FUNCTION_BLOCK "Select Station PB"   // FB45, SCL
{ S7_Optimized_Access := 'TRUE' }
VERSION : 0.1
   VAR_IN_OUT
      interface : "Push Button Data";
   END_VAR
   VAR
      "Get Button Feedback" : "Push Button: State Changes";
   END_VAR
   VAR_TEMP
      _interface : "Push Button Data";
      feedback : "Push Button Data: State Change Data";
   END_VAR
BEGIN
   REGION "BUFFER IN"
       #_interface := #interface;
   END_REGION

   REGION "PROCESS USER INPUT"
       #"Get Button Feedback"(interface := #_interface,
                              state_changes := #feedback);
   END_REGION

   REGION "ANIMATIONS"
       "Select Station PB: Private: Animations"(feedback := #feedback,
                                                interface := #_interface);
   END_REGION

   REGION "BUFFER OUT"
       #interface := #_interface;
   END_REGION
END_FUNCTION_BLOCK

FUNCTION "Select Station PB: Private: Animations" : Void   // FC94, SCL
{ S7_Optimized_Access := 'TRUE' }
VERSION : 0.1
   VAR_INPUT
      feedback : "Push Button Data: State Change Data";
   END_VAR
   VAR_IN_OUT
      interface : "Push Button Data";
   END_VAR
BEGIN
   REGION "COLOR"
       #interface.animate := "Bool.Animate"(true_color := "GREEN_LIGHT_BACKGROUND",
                                             false_color := "GRAY_BACKGROUND",
                                             evaluation_signal := #feedback.actuate.actual);
   END_REGION

   REGION "VISIBILITY"
       #interface.visible := TRUE;
   END_REGION

   REGION "ENABLED STATE"
       #interface.enable := TRUE;
   END_REGION
END_FUNCTION

// folder: Display: Warehouse/002 Settings/Select WIP Button

FUNCTION_BLOCK "Select WIP PB"   // FB46, SCL
{ S7_Optimized_Access := 'TRUE' }
VERSION : 0.1
   VAR_INPUT
      settings_meta : "Setting Meta Data";
      stations : "Station: All Stations";
   END_VAR
   VAR_IN_OUT
      interface : "Push Button Data";
   END_VAR
   VAR
      "Get Button Feedback" : "Push Button: State Changes";
   END_VAR
   VAR_TEMP
      _interface : "Push Button Data";
      enable : Bool;
      feedback : "Push Button Data: State Change Data";
      visible : Bool;
   END_VAR
BEGIN
   REGION "BUFFER IN"
       #_interface := #interface;
   END_REGION

   REGION "PROCESS USER INPUT"
       #"Get Button Feedback"(interface := #_interface,
                              state_changes := #feedback);
   END_REGION

   REGION "ANIMATIONS"
       "Select WIP PB: Private: Animations"(feedback := #feedback,
                                            settings_meta := #settings_meta,
                                            stations := #stations,
                                            interface := #_interface);
   END_REGION

   REGION "BUFFER OUT"
       #interface := #_interface;
   END_REGION
END_FUNCTION_BLOCK

FUNCTION "Select WIP PB: Private: Make Visible / Enable" : Bool   // FC92, SCL
{ S7_Optimized_Access := 'TRUE' }
VERSION : 0.1
   VAR_INPUT
      settings_meta : "Setting Meta Data";
      stations : "Station: All Stations";
   END_VAR
   VAR_TEMP
      ret : Bool;
      index_of_first_selected_station : Int;
      is_hmi_station : Bool;
      first_selected_station : "Station: Single Station";
      t_select_wip : "Push Button Data";
   END_VAR
BEGIN
   REGION "ARE SELECTED STATIONS HMI STATIONS?"
       #index_of_first_selected_station := "Get First Selected Station"(#settings_meta.selected_stations.stns);
       #first_selected_station := #stations.stn[#index_of_first_selected_station];
       #is_hmi_station := "Is_HMI_Station"(#first_selected_station);
   END_REGION

   REGION "HMI STATIONS"
       IF #is_hmi_station THEN
           #ret := TRUE;
       END_IF;
   END_REGION

   REGION "RETURN"
       #"Select WIP PB: Private: Make Visible / Enable" := #ret;
   END_REGION
END_FUNCTION

FUNCTION "Select WIP PB: Private: Animations" : Void   // FC123, SCL
{ S7_Optimized_Access := 'TRUE' }
VERSION : 0.1
   VAR_INPUT
      feedback : "Push Button Data: State Change Data";
      settings_meta : "Setting Meta Data";
      stations : "Station: All Stations";
   END_VAR
   VAR_IN_OUT
      interface : "Push Button Data";
   END_VAR
BEGIN
   REGION "COLOR"
       #interface.animate := "Bool.Animate"(true_color := "GREEN_LIGHT_BACKGROUND",
                                             false_color := "GRAY_BACKGROUND",
                                             evaluation_signal := #feedback.actuate.actual);
   END_REGION

   REGION "VISIBILITY"
       #interface.visible := "Select WIP PB: Private: Make Visible / Enable"(settings_meta := #settings_meta,
                                                                              stations := #stations);
   END_REGION

   REGION "ENABLED STATE"
       #interface.enable := "Select WIP PB: Private: Make Visible / Enable"(settings_meta := #settings_meta,
                                                                             stations := #stations);
   END_REGION
END_FUNCTION

// folder: Display: Warehouse/002 Settings/Selected WIP Table

FUNCTION_BLOCK "Selected_WIP_Table"   // FB30, SCL
{ S7_Optimized_Access := 'TRUE' }
VERSION : 0.1
   VAR_INPUT
      navigation_bar : "Nav Bar Data: PLC";
      pn_library : "Recipe: PN Text Library";
      saved_wips : "Recipe: HMI Stations Saved Wips";
      settings_meta : "Setting Meta Data";
      stations : "Station: All Stations";
      wip_library : "Recipe: Wip Text Library";
   END_VAR
   VAR_IN_OUT
      stationRows : Array[0..2] of "Settings Station Row Data";
   END_VAR
   VAR
      first_selected_station : Int;
      hmi_stations_selected : Bool;
      selected_stations : Array[0.."STATION_COUNT"] of Int;
      selected_list : "Selected_WIP_Table.Selected_Array";
      row_indices : Array[0..2] of DInt;
      inst_Table_Navigation : "Table Nav";
   END_VAR
   VAR_TEMP
      i : Int;
      p_stn : Int;
      wip_code : DInt;
      visible_rows : Int;
      first_null_index : DInt;
      _hmi_saved_station_index : Int;
      _wip_index : Int;
      _wip_module : "Station: Wip: Wip Module";
   END_VAR
   // row_indices[0] := 0;
   // row_indices[1] := 1;
   // row_indices[2] := 2;
BEGIN
   REGION "CLEAR OLD CONTENTS"    
       FOR #i := 0 TO 2 DO
           #stationRows[#i].line := "Cell_Data.Hide"();
           #stationRows[#i].dropzone := "Cell_Data.Hide"();
           #stationRows[#i].wip := "Cell_Data.Hide"();
           "Button_Row.Hide_Rows"(#stationRows[#i].btnRows);
       END_FOR;
   END_REGION


   REGION "EXIT ON NO SELECTED STATION"
       IF #settings_meta.selected_stations.count = 0 THEN
           RETURN;
       END_IF;
   END_REGION


   REGION "GET ARRAY OF SELECTED STATION INDICES"
       "Array.Int.Fill"(value := "NULL_TOKEN",
                        int_array := #selected_stations);
       "Selected_Stations.Indices"(selected_stations := #settings_meta.selected_stations,
                                   selected_stations_indices := #selected_stations);
       "Selected_WIP_Table.Build_List"(selected_stations := #selected_stations,
                                       selected_wips := #settings_meta.selected_wips.wips,
                                       selected_list := #selected_list);
   END_REGION


   REGION "DETERMINE IF SELECTED STATION IS AN HMI STATION"
       #first_selected_station := "Get First Selected Station"(#settings_meta.selected_stations.stns);
       #hmi_stations_selected := "Is_HMI_Station"(#stations.stn[#first_selected_station]);
   END_REGION


   REGION "TABLE DISPLAY POINTERS"
       #first_null_index := "Selected_WIP_Table.Selected_Array.First_Occurance"(selected_array := #selected_list,
                                                                                search_term := "NULL_TOKEN");
       #inst_Table_Navigation(first_null_index := #first_null_index,
                              tblData := #selected_list.me,
                              tblDisp := #stationRows,
                              tableNav := #navigation_bar,
                              rowIndices := #row_indices);
   END_REGION


   REGION "TABLE COMPONENTS"
       #visible_rows := DINT_TO_INT(#first_null_index) - 1;
       IF #visible_rows > 2 THEN
           #visible_rows := 2;
       END_IF;
       FOR #i := 0 TO #visible_rows DO
           #p_stn := #selected_list.me[#row_indices[#i]].station_pointer;
           #wip_code := #selected_list.me[#row_indices[#i]].wip_pointer;
           #stationRows[#i].line := "Selected_WIP_Table.Line_Label.Show"(station := #stations.stn[#p_stn]);
           #stationRows[#i].dropzone := "Selected_WIP_Table.Dropzone_Label.Show"(station := #stations.stn[#p_stn]);
           #stationRows[#i].wip := "Selected_WIP_Table.Wip_Label.Show"(wip_code := #wip_code,
                                                                       wip_library := #wip_library);
           #_wip_module := "Selected_WIP_Table.Get_WIP_Module"(stations := #stations,
                                                               saved_wips := #saved_wips,
                                                               station_pointer := #p_stn,
                                                               wip_code := #wip_code);
           "Button_Row.Show_Rows"(selected_butttons := #settings_meta.selected_btns,
                                  wip_module := #_wip_module,
                                  pn_library := #pn_library,
                                  button_rows := #stationRows[#i].btnRows);
       END_FOR;
   END_REGION
END_FUNCTION_BLOCK

FUNCTION "Selected_WIP_Table.Build_List" : Void   // FC219, SCL
{ S7_Optimized_Access := 'TRUE' }
VERSION : 0.1
   VAR_INPUT
      selected_stations : Array[*] of Int;
      selected_wips : Array[*] of DInt;
   END_VAR
   VAR_IN_OUT
      selected_list : "Selected_WIP_Table.Selected_Array";
   END_VAR
   VAR_TEMP
      _i : DInt;
      _j : DInt;
      _length : Struct
         stations : DInt;
         wips : DInt;
      END_STRUCT;
      _p : DInt;
   END_VAR
BEGIN
   REGION "PREPARE ARRAY"
       "Selected_WIP_Table.Selected_Array.Fill"(token := -1,
                                                selected_list := #selected_list);
   END_REGION


   REGION "GET UPPER LIMIT FOR OUTER LOOP"
       #_length.stations := "Array.Int.First_Occurance"(int_array := #selected_stations,
                                                        search_term := "NULL_TOKEN");
       #_length.stations -= 1;
       #_length.stations := "DInt.Clip.Minimum"(value := #_length.stations,
                                                minimum := 0);
   END_REGION


   REGION "GET LIMIT FOR INNER LOOP"
       #_length.wips := "Array.DInt.First_Occurance"(dint_array := #selected_wips,
                                                     search_term := "NULL_TOKEN");
       #_length.wips -= 1;
       #_length.wips := "DInt.Clip.Minimum"(value := #_length.wips,
                                            minimum := 0);
   END_REGION


   REGION "BUILD ARRAY"
       FOR #_i := 0 TO #_length.stations DO
           FOR #_j := 0 TO #_length.wips DO
               #_p := #_i * (#_length.wips + 1) + #_j;
               #selected_list.me[#_p].station_pointer := #selected_stations[#_i];
               #selected_list.me[#_p].wip_pointer := #selected_wips[#_j];
           END_FOR;
       END_FOR;
   END_REGION
END_FUNCTION

FUNCTION "Selected_WIP_Table.Selected_Array.Fill" : Void   // FC221, SCL
{ S7_Optimized_Access := 'TRUE' }
VERSION : 0.1
   VAR_INPUT
      token : Int;
   END_VAR
   VAR_IN_OUT
      selected_list : "Selected_WIP_Table.Selected_Array";
   END_VAR
   VAR_TEMP
      _i : DInt;
      _length : DInt;
   END_VAR
BEGIN
   #_length := UDINT_TO_DINT("Array.Any.Length"(#selected_list.me));
   #_length -= 1;

   FOR #_i := 0 TO #_length DO
       #selected_list.me[#_i].station_pointer := #token;
       #selected_list.me[#_i].wip_pointer := INT_TO_DINT(#token);
   END_FOR;
END_FUNCTION

FUNCTION "Selected_WIP_Table.Selected_Array.Is_Element" : Bool   // FC228, SCL
{ S7_Optimized_Access := 'TRUE' }
VERSION : 0.1
   VAR_INPUT
      selected_array : "Selected_WIP_Table.Selected_Array";
      search_term : Int;
   END_VAR
   VAR_TEMP
      _i : DInt;
      _length : DInt;
   END_VAR
BEGIN
   REGION "LOCAL VARIABLES"
       #_length := UDINT_TO_DINT("Array.Any.Length"(#selected_array.me)) - 1;
   END_REGION


   REGION "SEARCH ARRAY"
       FOR #_i := 0 TO #_length DO
           IF #selected_array.me[#_i].station_pointer <> #search_term THEN
               CONTINUE;
           END_IF;
           #"Selected_WIP_Table.Selected_Array.Is_Element" := TRUE;
           RETURN;
       END_FOR;
   END_REGION


   REGION "NOT FOUND"
       #"Selected_WIP_Table.Selected_Array.Is_Element" := FALSE;
       RETURN;
   END_REGION
END_FUNCTION

FUNCTION "Selected_WIP_Table.Selected_Array.First_Occurance" : DInt   // FC229, SCL
{ S7_Optimized_Access := 'TRUE' }
VERSION : 0.1
   VAR_INPUT
      selected_array : "Selected_WIP_Table.Selected_Array";
      search_term : Int;
   END_VAR
   VAR_TEMP
      _i : DInt;
      _length : UDInt;
   END_VAR
BEGIN
   REGION "NOTES"
       (* 
       This function returns the first occurance of the search term.
       This function meant for use with collapsed arrays.
       See "Array.Int.Collapse" for collapse functionality.
       *)
   END_REGION


   REGION "GET LENGTH OF INPUT ARRAY"
       #_length := "Array.Any.Length"(#selected_array.me);
   END_REGION


   REGION "FIND FIRST SEARCH TERM, -1 IF NONE"
       (*
       Its worth noting that "Array.Int.Is_Element" could return the index of the search term
       as an output, saving the processor some work. 
       The rework is justified by increased encapsulation.
       The time complexity for "Array.Int.First_Occurance" remains O(n).
       *)
       IF NOT "Selected_WIP_Table.Selected_Array.Is_Element"(selected_array:=#selected_array, search_term:=#search_term) THEN
           #"Selected_WIP_Table.Selected_Array.First_Occurance" := -1;
           RETURN;
       END_IF;
       WHILE #selected_array.me[#_i].station_pointer <> #search_term AND DINT_TO_UDINT(#_i) < #_length DO
           #_i += 1;
       END_WHILE;
   END_REGION


   REGION "SEARCH TERM FOUND"
       #"Selected_WIP_Table.Selected_Array.First_Occurance" := #_i;
       RETURN;
   END_REGION
END_FUNCTION

FUNCTION "Selected_WIP_Table.Get_WIP_Module" : "Station: Wip: Wip Module"   // FC234, SCL
{ S7_Optimized_Access := 'TRUE' }
VERSION : 0.1
   VAR_INPUT
      stations : "Station: All Stations";
      saved_wips : "Recipe: HMI Stations Saved Wips";
      station_pointer : Int;
      wip_code : DInt;
   END_VAR
   VAR_TEMP
      _hmi_station_pointer : Int;
      _wip_pointer : Int;
   END_VAR
BEGIN
   IF #wip_code = "NULL_TOKEN" THEN
       #"Selected_WIP_Table.Get_WIP_Module" := #stations.stn[#station_pointer].wipCmpts;
       RETURN;
   END_IF;

   #_hmi_station_pointer := "WIP.Global_Index_to_HMI_Station_Index"(global_index := #station_pointer,
                                                                    saved_WIPs := #saved_wips);

   #_wip_pointer := "WIP.Code_to_Index"(saved_wip := #saved_wips.stn[#_hmi_station_pointer],
                                        wip_code := #wip_code);

   #"Selected_WIP_Table.Get_WIP_Module" := #saved_wips.stn[#_hmi_station_pointer].wip[#_wip_pointer];
   RETURN;
END_FUNCTION

// folder: Display: Warehouse/002 Settings/Selected WIP Table/Button Row

FUNCTION "Button_Row.Hide" : "Settings Station Row Button Row Data"   // FC210, SCL
{ S7_Optimized_Access := 'TRUE' }
VERSION : 0.1
   VAR_TEMP
      _ret : "Settings Station Row Button Row Data";
   END_VAR
BEGIN
   #_ret.button := "Cell_Data.Hide"();
   #_ret.total := "Cell_Data.Hide"();
   #_ret.critical := "Cell_Data.Hide"();
   #_ret.singlePN := "Cell_Data.Hide"();
   #_ret.doublePN := "Cell_Data.Hide"();
   #"Button_Row.Hide" := #_ret;
END_FUNCTION

FUNCTION "Button_Row.Hide_Rows" : Void   // FC211, SCL
{ S7_Optimized_Access := 'TRUE' }
VERSION : 0.1
   VAR_IN_OUT
      button_rows : Array[*] of "Settings Station Row Button Row Data";
   END_VAR
   VAR_TEMP
      _i : Int;
   END_VAR
BEGIN
   FOR #_i := 0 TO UDINT_TO_INT("Array.Any.Length"(#button_rows)) - 1 DO
       #button_rows[#_i] := "Button_Row.Hide"();
   END_FOR;
END_FUNCTION

FUNCTION "Button_Row.Show" : "Settings Station Row Button Row Data"   // FC212, SCL
{ S7_Optimized_Access := 'TRUE' }
VERSION : 0.1
   VAR_INPUT
      button_number : Int;
      selected : Bool;
      pn_library : "Recipe: PN Text Library";
      wip_module : "Station: Wip: Wip Module";
   END_VAR
   VAR_TEMP
      _return : "Settings Station Row Button Row Data";
      _pn : "Cell Data";
   END_VAR
BEGIN
   #_return.button := "Button_Row.Button_Label.Show"(button_number := #button_number,
                                                     selected := #selected);

   #_return.total := "Button_Row.Total.Show"(selected := #selected,
                                             button_number := #button_number,
                                             wip_module := #wip_module);

   #_return.critical := "Button_Row.Critical.Show"(button_number := #button_number,
                                                   selected := #selected,
                                                   wip_module := #wip_module);

   #_pn := "Button_Row.Part_Number.Show"(button_number := #button_number,
                                         pn_library := #pn_library,
                                         selected := #selected,
                                         wip_module := #wip_module);

   IF "Part_Number.Is_Single"(#wip_module.pnCode[#button_number]) THEN
       #_return.singlePN := #_pn;
   END_IF;
   IF "Part_Number.Is_Double"(#wip_module.pnCode[#button_number]) THEN
       #_return.doublePN := #_pn;
   END_IF;
   #"Button_Row.Show" := #_return;
END_FUNCTION

FUNCTION "Button_Row.Show_Rows" : Void   // FC218, SCL
{ S7_Optimized_Access := 'TRUE' }
VERSION : 0.1
   VAR_INPUT
      selected_butttons : "Selected Buttons";
      wip_module : "Station: Wip: Wip Module";
      pn_library : "Recipe: PN Text Library";
   END_VAR
   VAR_IN_OUT
      button_rows : Array[*] of "Settings Station Row Button Row Data";
   END_VAR
   VAR_TEMP
      _i : Int;
      _remap : Int;
   END_VAR
BEGIN
   FOR #_i := 0 TO UDINT_TO_INT("Array.Any.Length"(#button_rows)) - 1 DO
       #_remap := "KP8.DURL_to_LRUD"(#_i);
       #button_rows[#_i] := "Button_Row.Show"(button_number := #_remap,
                                              selected := #selected_butttons.btns[#_i],
                                              pn_library := #pn_library,
                                              wip_module := #wip_module);
   END_FOR;
END_FUNCTION

// folder: Display: Warehouse/002 Settings/Selected WIP Table/Button Row/Single Button

FUNCTION "Button_Row.Button_Label.Show" : "Cell Data"   // FC213, SCL
{ S7_Optimized_Access := 'TRUE' }
VERSION : 0.1
   VAR_INPUT
      button_number : Int;
      selected : Bool;
   END_VAR
   VAR_TEMP
      _animate : Int;
      _data : WString;
   END_VAR
BEGIN
   #_animate := "Bool.Animate"(true_color := "BLUE_LIGHT_BACKGROUND",
                               false_color := "GRAY_BACKGROUND",
                               evaluation_signal := #selected);
   #_data := "Trim"("Strip Sign"(INT_TO_WSTRING(#button_number)));
   #"Button_Row.Button_Label.Show" := "Cell_Data.Show"(animate := #_animate, data := #_data);
END_FUNCTION

FUNCTION "Button_Row.Total.Show" : "Cell Data"   // FC214, SCL
{ S7_Optimized_Access := 'TRUE' }
VERSION : 0.1
   VAR_INPUT
      button_number : Int;
      selected : Bool;
      wip_module : "Station: Wip: Wip Module";
   END_VAR
   VAR_TEMP
      _animation : Int;
      _data : WString;
   END_VAR
BEGIN
   #_animation := "Bool.Animate"(true_color := "BLUE_LIGHT_BACKGROUND",
                                 false_color := "GRAY_BACKGROUND",
                                 evaluation_signal := #selected);

   #_data := "Button_Row.Total.Extract_String"(button_number := #button_number,
                                               wip_module := #wip_module);

   #"Button_Row.Total.Show" := "Cell_Data.Show"(animate := #_animation,
                                                data := #_data);
END_FUNCTION

FUNCTION "Button_Row.Critical.Show" : "Cell Data"   // FC215, SCL
{ S7_Optimized_Access := 'TRUE' }
VERSION : 0.1
   VAR_INPUT
      button_number : Int;
      selected : Bool;
      wip_module : "Station: Wip: Wip Module";
   END_VAR
   VAR_TEMP
      _animate : Int;
      _data : WString;
   END_VAR
BEGIN
   #_animate := "Bool.Animate"(true_color := "BLUE_LIGHT_BACKGROUND",
                               false_color := "GRAY_BACKGROUND",
                               evaluation_signal := #selected);

   #_data := "Button_Row.Critical.Extract_String"(button_number := #button_number,
                                                  wip_module := #wip_module);

   #"Button_Row.Critical.Show" := "Cell_Data.Show"(animate := #_animate, data := #_data);
END_FUNCTION

FUNCTION "Button_Row.Part_Number.Show" : "Cell Data"   // FC217, SCL
{ S7_Optimized_Access := 'TRUE' }
VERSION : 0.1
   VAR_INPUT
      button_number : Int;
      pn_library : "Recipe: PN Text Library";
      selected : Bool;
      wip_module : "Station: Wip: Wip Module";
   END_VAR
   VAR_TEMP
      _animation : Int;
      _data : WString;
      _pn_code : DInt;
   END_VAR
BEGIN
   #_animation := "Bool.Animate"(true_color := "BLUE_LIGHT_BACKGROUND",
                                 false_color := "GRAY_BACKGROUND",
                                 evaluation_signal := #selected);

   #_pn_code := "Button_Row.Part_Number.Extract_Code"(button_number := #button_number,
                                                      wip_module := #wip_module);

   #_data := "Part_Number.Code_to_WString"(pnLib := #pn_library,
                                           pnCode := #_pn_code);

   #"Button_Row.Part_Number.Show" := "Cell_Data.Show"(animate := #_animation,
                                                      data := #_data);
END_FUNCTION

FUNCTION "Button_Row.Total.Extract_String" : WString   // FC230, SCL
{ S7_Optimized_Access := 'TRUE' }
VERSION : 0.1
   VAR_INPUT
      button_number : Int;
      wip_module : "Station: Wip: Wip Module";
   END_VAR
BEGIN
   #"Button_Row.Total.Extract_String" := "Timer.Real_to_WString"(#wip_module.timers.ptAllotted[#button_number]);
   RETURN;
END_FUNCTION

FUNCTION "Button_Row.Part_Number.Extract_Code" : DInt   // FC231, SCL
{ S7_Optimized_Access := 'TRUE' }
VERSION : 0.1
   VAR_INPUT
      button_number : Int;
      wip_module : "Station: Wip: Wip Module";
   END_VAR
   VAR_TEMP
      _hmi_station_pointer : Int;
      _pn_code : DInt;
      _wip_pointer : Int;
   END_VAR
BEGIN
   #"Button_Row.Part_Number.Extract_Code" := #wip_module.pnCode[#button_number];
   RETURN;
END_FUNCTION

FUNCTION "Button_Row.Critical.Extract_String" : WString   // FC232, SCL
{ S7_Optimized_Access := 'TRUE' }
VERSION : 0.1
   VAR_INPUT
      button_number : Int;
      wip_module : "Station: Wip: Wip Module";
   END_VAR
BEGIN
   #"Button_Row.Critical.Extract_String" := "Timer.Real_to_WString"(#wip_module.timers.ptCritical[#button_number]);
   RETURN;
END_FUNCTION

// folder: Display: Warehouse/002 Settings/Selected WIP Table/Dropzone Label

FUNCTION "Selected_WIP_Table.Dropzone_Label.Show" : "Cell Data"   // FC200, SCL
{ S7_Optimized_Access := 'TRUE' }
VERSION : 0.1
   VAR_INPUT
      station : "Station: Single Station";
   END_VAR
BEGIN
   #"Selected_WIP_Table.Dropzone_Label.Show" := "Cell_Data.Show"(animate := "GRAY_BACKGROUND",
                                                                 data := "Trim"("Strip Sign"(USINT_TO_WSTRING(#station.id.dropZone))));
END_FUNCTION

// folder: Display: Warehouse/002 Settings/Selected WIP Table/Line Label

FUNCTION "Selected_WIP_Table.Line_Label.Show" : "Cell Data"   // FC199, SCL
{ S7_Optimized_Access := 'TRUE' }
VERSION : 0.1
   VAR_INPUT
      station : "Station: Single Station";
   END_VAR
   VAR CONSTANT
      SHOW : Bool := TRUE;
   END_VAR
BEGIN
   #"Selected_WIP_Table.Line_Label.Show" := "Cell_Data.Show"(animate := "GRAY_BACKGROUND",
                                                             data := #station.id.lineName);
END_FUNCTION

// folder: Display: Warehouse/002 Settings/Selected WIP Table/Wip Label

FUNCTION "Selected_WIP_Table.Wip_Label.Show" : "Cell Data"   // FC201, SCL
{ S7_Optimized_Access := 'TRUE' }
VERSION : 0.1
   VAR_INPUT
      wip_code : DInt;
      wip_library : "Recipe: Wip Text Library";
   END_VAR
   VAR_TEMP
      _delimeters : Array[0..9] of WString[1];
      _data : WString;
   END_VAR
   VAR CONSTANT
      SHOW : Bool := TRUE;
   END_VAR
BEGIN
   IF #wip_code = "NULL_TOKEN" THEN
       #"Selected_WIP_Table.Wip_Label.Show" := "Cell_Data.Hide"();
       RETURN;
   END_IF;

   #_data := "WIP.Code_to_WString"(wipTxtLib := #wip_library,
                                   code := #wip_code);
   #_delimeters[0] := WSTRING#' ';
   #_delimeters[1] := WSTRING#'-';
   #_delimeters[2] := WSTRING#'.';
   #_data := "WString.Word_Wrap"(delimeters := #_delimeters,
                                 line_length := 20,
                                 wstring_in := #_data);

   #"Selected_WIP_Table.Wip_Label.Show" := "Cell_Data.Show"(animate := "GRAY_BACKGROUND", data := #_data);
END_FUNCTION

// folder: Display: Warehouse/002 Settings/Total IO Field

FUNCTION_BLOCK "Total_IO_Field"   // FB49, SCL
{ S7_Optimized_Access := 'TRUE' }
VERSION : 0.1
   VAR_INPUT
      settings_meta : "Setting Meta Data";
      stations : "Station: All Stations";
   END_VAR
   VAR_IN_OUT
      interface : "IO Field Data: Label with Data";
      state_changes : "State Changes: Real";
   END_VAR
   VAR
      Total_IO_Field : "IO Field: State Changes";
      Detect_State_Changes : "Real.State_Change";
   END_VAR
   VAR_TEMP
      _interface : "IO Field Data: Label with Data";
      feedback : "IO Field: State Change Data";
   END_VAR
BEGIN
   REGION "BUFFER IN"
       #_interface := #interface;
   END_REGION

   REGION "PROCESS USER INPUT"
       #Total_IO_Field(interface := #_interface,
                       feedback := #feedback);
       #Detect_State_Changes(value := "Timer.WString_to_Real"(#interface.value),
                             get_real := #state_changes);
   END_REGION

   REGION "BUFFER OUT"
       "Total_IO_Field.Animate"(feedback := #feedback,
                                settings_meta := #settings_meta,
                                stations := #stations,
                                interface := #_interface);
   END_REGION

   REGION "BUFFER OUT"
       #interface := #_interface;
   END_REGION
END_FUNCTION_BLOCK

FUNCTION "Total_IO_Field.Make_Visible_Enable" : Bool   // FC189, SCL
{ S7_Optimized_Access := 'TRUE' }
VERSION : 0.1
   VAR_INPUT
      setting_meta : "Setting Meta Data";
   END_VAR
BEGIN
   #"Total_IO_Field.Make_Visible_Enable" := #setting_meta.selected_btns.count > 0;
END_FUNCTION

FUNCTION "Total_IO_Field.Animate" : Void   // FC190, SCL
{ S7_Optimized_Access := 'TRUE' }
VERSION : 0.1
   VAR_INPUT
      feedback : "IO Field: State Change Data";
      settings_meta : "Setting Meta Data";
      stations : "Station: All Stations";
   END_VAR
   VAR_IN_OUT
      interface : "IO Field Data: Label with Data";
   END_VAR
   VAR_TEMP
      _visible_enabled : Bool;
   END_VAR
BEGIN
   REGION "COLOR"
   #interface.animate := "WHITE_BACKGROUND";
   END_REGION


   REGION "SET STATE"
       #_visible_enabled := "Total_IO_Field.Make_Visible_Enable"(setting_meta := #settings_meta);
   END_REGION


   REGION "VISIBILITY
       #interface.visible := #_visible_enabled;
   END_REGION


   REGION "ENABLE"
       #interface.enable := #_visible_enabled;
   END_REGION


   REGION "POPULATE VALUE"
       IF #settings_meta.button_selection_change.selection_change THEN
           #interface.value := "Total_IO_Field.Populate_Value"(hidden := NOT #_visible_enabled,
                                                               selected_buttons := #settings_meta.selected_btns,
                                                               selected_stations := #settings_meta.selected_stations,
                                                               stations := #stations);
       END_IF;
   END_REGION
END_FUNCTION

FUNCTION "Total_IO_Field.Populate_Value" : WString   // FC292, SCL
{ S7_Optimized_Access := 'TRUE' }
VERSION : 0.1
   VAR_INPUT
      hidden : Bool;
      selected_buttons : "Selected Buttons";
      selected_stations : "Selected Stations";
      stations : "Station: All Stations";
   END_VAR
   VAR_TEMP
      _critical : WString;
      _p_station : Int;
      _p_button : Int;
   END_VAR
   VAR CONSTANT
      BLANK : WString;
      ZERO : WChar := WCHAR#'0';
   END_VAR
BEGIN
   IF #hidden THEN
       #"Total_IO_Field.Populate_Value" := #BLANK;
       RETURN;
   END_IF;
   #_p_station := "Selected_Stations.Get_First_Selected_Station"(#selected_stations);
   #_p_button := "Selected_Buttons.Get_First_Selected_Button"(#selected_buttons);
   #_critical := "Timer.Real_to_WString"(#stations.stn[#_p_station].wipCmpts.timers.ptAllotted[#_p_button]);
   #"Total_IO_Field.Populate_Value" := #_critical;
END_FUNCTION

// folder: Display: Warehouse/Pop Ups/Pop Up Utilities

FUNCTION "Animate Array: PB Data Activation" : Bool   // FC95, SCL
{ S7_Optimized_Access := 'TRUE' }
VERSION : 0.1
   VAR_INPUT
      element_index : Int;
      visible_element_count : Int;
   END_VAR
   VAR_TEMP
      ret : Bool;
   END_VAR
BEGIN
   REGION "TURN ON A NUMBER OF BUTTONS EQUAL TO THE NUMBER OF STATIONS"
       IF #element_index < #visible_element_count THEN
           #ret := TRUE;
       END_IF;
       IF #element_index >= #visible_element_count THEN
           #ret := FALSE;
       END_IF;
   END_REGION

   REGION "RETURN"
       #"Animate Array: PB Data Activation" := #ret;
   END_REGION
END_FUNCTION

FUNCTION "Pop Up: Nav Bar: Button Animation" : Void   // FC97, SCL
{ S7_Optimized_Access := 'TRUE' }
VERSION : 0.1
   VAR_INPUT
      selectable_elements : Int;
      visible_rows : Int;
   END_VAR
   VAR_IN_OUT
      button : "Push Button Data";
   END_VAR
   VAR_TEMP
      ret : "Push Button Data";
   END_VAR
BEGIN
   REGION "SHOW NAV BAR"
       IF #selectable_elements > #visible_rows THEN

           REGION "GET CURRENT STATE FOR PRESS"
               #ret := #button;
           END_REGION

           REGION "ANIMATION"
               #ret.animate := "Bool.Animate"(true_color := "GREEN_LIGHT_BACKGROUND",
                                              false_color := "GRAY_BACKGROUND",
                                              evaluation_signal := #button.actuate);
           END_REGION

           REGION "ENABLE"
               #ret.enable := TRUE;
           END_REGION

           REGION "LIST SELECT"
               #ret.listSelect := 0;
           END_REGION

           REGION "VISIBLE"
               #ret.visible := TRUE;
           END_REGION

       END_IF;
   END_REGION


   REGION "HIDE NAV BAR"
       IF #selectable_elements <= #visible_rows THEN

           REGION "DIABLE"
               #ret.enable := FALSE;
           END_REGION

           REGION "INVISIBLE"
               #ret.visible := FALSE;
           END_REGION

       END_IF;
   END_REGION


   REGION "RETURN"
       #button := #ret;
   END_REGION
END_FUNCTION

FUNCTION "Pop Up: Map Select Button Actuations" : Void   // FC117, SCL
{ S7_Optimized_Access := 'TRUE' }
VERSION : 0.1
   VAR_INPUT
      screen_elements : Variant;
   END_VAR
   VAR_IN_OUT
      actuations_as_ints : Variant;
   END_VAR
   VAR_TEMP
      i : Int;
      len_udint : UDInt;
      len_int : Int;
      ret : Array[0..#u_bound_simple] of Int;
      status : Int;
      t_select_btns : Array[0..#u_bound_complex] of "Push Button Data";
   END_VAR
   VAR CONSTANT
      u_bound_simple : Int := 99;
      u_bound_complex : Int := 29;
   END_VAR
BEGIN
   REGION "GET PARAMETERS"
       #len_udint := CountOfElements(#screen_elements);
       #len_int := UDINT_TO_INT(#len_udint) - 1;
   END_REGION

   REGION "COPY TO LOCAL"
       #status := MOVE_BLK_VARIANT(SRC := #screen_elements,
                                   COUNT := #len_udint,
                                   SRC_INDEX := 0,
                                   DEST_INDEX := 0,
                                   DEST => #t_select_btns);
   END_REGION

   REGION "MAP ACTUATIONS"    
       FOR #i := 0 TO #len_int DO
           IF #t_select_btns[#i].actuate THEN
               #ret[#i] := 1;
           END_IF;
       END_FOR;
   END_REGION

   REGION "RETURN"
       #status := MOVE_BLK_VARIANT(SRC := #ret,
                                   COUNT := #len_udint,
                                   SRC_INDEX := 0,
                                   DEST_INDEX := 0,
                                   DEST => #actuations_as_ints);
   END_REGION
END_FUNCTION

FUNCTION "Pop Up: Nav Bar: Animate" : Void   // FC135, SCL
{ S7_Optimized_Access := 'TRUE' }
VERSION : 0.1
   VAR_INPUT
      selectable_element_count : Int;
      visible_rows : Int;
   END_VAR
   VAR_IN_OUT
      nav_bar : "Nav Bar Data";
   END_VAR
BEGIN
       REGION "NOTES"
           // mapping is necessary because hmi faceplate data structures
           // cannot consist of embedded udts
       END_REGION

       REGION "MAP HMI TO PLC"
           "NavBar: Map HMI to PLC"(hmi := #nav_bar.hmi,
                                          plc := #nav_bar.plc);
       END_REGION

       REGION "ANIMATION CALLS"
           "Pop Up: Nav Bar: Button Animation"(selectable_elements := #selectable_element_count,
                                               visible_rows := #visible_rows,
                                               button := #nav_bar.plc.top);
           "Pop Up: Nav Bar: Button Animation"(selectable_elements := #selectable_element_count,
                                               visible_rows := #visible_rows,
                                               button := #nav_bar.plc.pageUp);
           "Pop Up: Nav Bar: Button Animation"(selectable_elements := #selectable_element_count,
                                               visible_rows := #visible_rows,
                                               button := #nav_bar.plc.lineUp);
           "Pop Up: Nav Bar: Button Animation"(selectable_elements := #selectable_element_count,
                                               visible_rows := #visible_rows,
                                               button := #nav_bar.plc.lineDown);
           "Pop Up: Nav Bar: Button Animation"(selectable_elements := #selectable_element_count,
                                               visible_rows := #visible_rows,
                                               button := #nav_bar.plc.pageDown);
           "Pop Up: Nav Bar: Button Animation"(selectable_elements := #selectable_element_count,
                                               visible_rows := #visible_rows,
                                               button := #nav_bar.plc.bottom);
       END_REGION

       REGION "MAP PLC TO HMI"
           "NavBar: Map PLC to HMI"(plc := #nav_bar.plc,
                                          hmi := #nav_bar.hmi);
       END_REGION
END_FUNCTION

FUNCTION "Clear WIP Selection Meta Data" : Void   // FC193, SCL
{ S7_Optimized_Access := 'TRUE' }
VERSION : 0.1
   VAR_IN_OUT
      selected_wips : "Selected Wips";
   END_VAR
   VAR_TEMP
      i : Int;
      selected_wips_array : Array[0.."WIP_COUNT"] of DInt;
   END_VAR
BEGIN
   "Array.DInt.Fill"(int_in := INT_TO_DINT("NULL_TOKEN"),
                     array_out => #selected_wips.wips);
   #selected_wips.count := 0;
END_FUNCTION

FUNCTION "Clear Button Selection Meta Data" : Void   // FC194, SCL
{ S7_Optimized_Access := 'TRUE' }
VERSION : 0.1
   VAR_IN_OUT
      selected_buttons : "Selected Buttons";
   END_VAR
   VAR_TEMP
      i : Int;
   END_VAR
BEGIN
   #selected_buttons.count := 0;
   FOR #i := 0 TO "BUTTON_COUNT" DO
       #selected_buttons.btns[#i] := FALSE;
   END_FOR;
END_FUNCTION

// folder: Display: Warehouse/Pop Ups/Select Buttons

FUNCTION_BLOCK "Pop Up: Select Buttons"   // FB25, SCL
{ S7_Optimized_Access := 'TRUE' }
VERSION : 0.1
   VAR_IN_OUT
      interface : "Select Button";
      selected_buttons : "Selected Buttons";
      meta_data : "Setting Meta Data";
   END_VAR
   VAR
      "inst Pop Up: Select Buttons: Select Buttons" : "Pop Up: Select Buttons: Select Buttons";
      Button_Selection_Change : "Selected_Buttons.Selection_Change";
   END_VAR
BEGIN
   REGION "ANIMATION"
       "Pop Up: Select Buttons: Animations"(interface := #interface,
                                            selected := #selected_buttons);
   END_REGION


   REGION "PERFORM BUTTON SELECTION"
       #"inst Pop Up: Select Buttons: Select Buttons"(interface := #interface,
                                                      selected_buttons := #selected_buttons);
   END_REGION


   REGION "CHECK FOR BUTTON SELECTION CHANGE"
       #Button_Selection_Change(selected_buttons := #selected_buttons,
                                selection_change := #meta_data.button_selection_change);
   END_REGION


   REGION "HOUSE KEEPING FOR STATION SELECTION CHANGE"
       IF #meta_data.station_selection_change.selection_change THEN
           "Clear Button Selection Meta Data"(#meta_data.selected_btns);
       END_IF;
   END_REGION
END_FUNCTION_BLOCK

FUNCTION_BLOCK "Pop Up: Select Buttons: Select Buttons"   // FB27, SCL
{ S7_Optimized_Access := 'TRUE' }
VERSION : 0.1
   VAR_IN_OUT
      interface : "Select Button";
      selected_buttons : "Selected Buttons";
   END_VAR
   VAR
      "inst Pulses: Button Collection" : "Pulses: Button Collection";
   END_VAR
   VAR_TEMP
      actuation_pulses : Array[0.."BUTTON_COUNT"] of Bool;
      actuations_as_ints : Array[0.."BUTTON_COUNT"] of Int;
      i : Int;
      pulses_as_ints : Array[0.."BUTTON_COUNT"] of Int;
   END_VAR
BEGIN
   "Pop Up: Map Select Button Actuations"(screen_elements := #interface.buttons,
                                          actuations_as_ints := #actuations_as_ints);
   #"inst Pulses: Button Collection"(btns := #actuations_as_ints,
                                     pulses := #pulses_as_ints);
   "Pop Up: Select Buttons: Pulse Ints to Bools"(pulses_as_ints := #pulses_as_ints,
                                                 pulses_as_bools => #actuation_pulses);
   FOR #i := 0 TO "BUTTON_COUNT" DO
       "Toggle"(pulse := #actuation_pulses[#i],
                state := #selected_buttons.btns[#i]);
   END_FOR;
   #selected_buttons.count := "Count Selected Buttons"(#selected_buttons.btns);
END_FUNCTION_BLOCK

FUNCTION_BLOCK "Selected_Buttons.Selection_Change"   // FB59, SCL
{ S7_Optimized_Access := 'TRUE' }
VERSION : 0.1
   VAR_INPUT
      selected_buttons : "Selected Buttons";
   END_VAR
   VAR_IN_OUT
      selection_change : "Selected_Buttons.Selection_Change.UDT";
   END_VAR
   VAR
      old : Struct
         selected_buttons : "Selected Buttons";
      END_STRUCT;
   END_VAR
   VAR_TEMP
      _i : Int;
      _return : "Selected_Buttons.Selection_Change.UDT";
   END_VAR
BEGIN
   REGION "SCAN FOR CHANGE"
       FOR #_i := 0 TO "BUTTON_COUNT" DO
           IF #selected_buttons.btns[#_i] <> #old.selected_buttons.btns[#_i] THEN
               #_return.selection_change := TRUE;
               #_return.button_index := #_i;
               IF #selected_buttons.btns[#_i] AND NOT #old.selected_buttons.btns[#_i] THEN
                   #_return.rising := TRUE;
                   #_return.falling := FALSE;
               END_IF;
               IF NOT #selected_buttons.btns[#_i] AND #old.selected_buttons.btns[#_i] THEN
                   #_return.rising := FALSE;
                   #_return.falling := TRUE;
               END_IF;
               EXIT;
           END_IF;
       END_FOR;
   END_REGION


   REGION "SAVE TO OLD"
       #old.selected_buttons := #selected_buttons;
   END_REGION


   REGION "RETURN"
       #selection_change := #_return;
   END_REGION
END_FUNCTION_BLOCK

FUNCTION "Pop Up: Select Buttons: Animations" : Void   // FC116, SCL
{ S7_Optimized_Access := 'TRUE' }
VERSION : 0.1
   VAR_IN_OUT
      interface : "Select Button";
      selected : "Selected Buttons";
   END_VAR
   VAR_TEMP
      i : Int;
      selected_stations_count : Int;
      t_interface : "Select Button";
   END_VAR
BEGIN
   REGION "COPY TO LOCAL"
       #t_interface := #interface;
   END_REGION

   REGION "CLOSE POPUP BUTTON"
       #t_interface.close_screen.animate := "Bool.Animate"(true_color := "GREEN_LIGHT_BACKGROUND",
                                                           false_color := "RED_LIGHT_BACKGROUND",
                                                           evaluation_signal := #interface.close_screen.actuate);
   END_REGION


   REGION "BUTTON SELECTION BUTTONS"
       FOR #i := 0 TO "BUTTON_COUNT" DO
           #t_interface.buttons[#i].animate := "Bool.Animate"(true_color := "GREEN_LIGHT_BACKGROUND",
                                                              false_color := "GRAY_BACKGROUND",
                                                              evaluation_signal := #interface.buttons[#i].actuate);
           #t_interface.buttons[#i].enable := TRUE;
           #t_interface.buttons[#i].visible := TRUE;
           IF #selected.btns[#i] THEN
               #t_interface.buttons[#i].animate := "BLUE_LIGHT_BACKGROUND";
           END_IF;
       END_FOR;
   END_REGION


   REGION "DRAW"
       #interface := #t_interface;
   END_REGION
END_FUNCTION

FUNCTION "Pop Up: Select Buttons: Pulse Ints to Bools" : Void   // FC118, SCL
{ S7_Optimized_Access := 'TRUE' }
VERSION : 0.1
   VAR_INPUT
      pulses_as_ints : Array[0.."BUTTON_COUNT"] of Int;
   END_VAR
   VAR_OUTPUT
      pulses_as_bools : Array[0.."BUTTON_COUNT"] of Bool;
   END_VAR
   VAR_TEMP
      i : Int;
      ret : Array[0.."BUTTON_COUNT"] of Bool;
   END_VAR
BEGIN
   REGION "MAP TO BOOLS"
       FOR #i := 0 TO "BUTTON_COUNT" DO
           #ret[#i] := #pulses_as_ints[#i].%X0;
       END_FOR;
   END_REGION

   REGION "RETURN"
       #pulses_as_bools := #ret;
   END_REGION
END_FUNCTION

// folder: Display: Warehouse/Pop Ups/Select Station

FUNCTION_BLOCK "Pop Up: Select Stations"   // FB21, SCL
{ S7_Optimized_Access := 'TRUE' }
VERSION : 0.1
   VAR_INPUT
      all_stations : "Station: All Stations";
      saved_WIPs : "Recipe: HMI Stations Saved Wips";
   END_VAR
   VAR_IN_OUT
      interface : "Select Station";
      meta_data : "Setting Meta Data";
   END_VAR
   VAR
      "inst Patch for Table Nav in Select Station Popup" : "Patch for Table Nav in Select Station Popup";
      "inst Select Station Button Pulses" : "Pulses: Button Collection";
      "inst Selection Change" : "Selected_Stations.Selection_Change";
      "inst Table Nav" : "Table Nav";
      vis_stns_as_dint : Array[0.."_SELECT_STATION_BUTTON_COUNT"] of DInt;
      visable_stns : Array[0.."_SELECT_STATION_BUTTON_COUNT"] of Int;
   END_VAR
   VAR_TEMP
      actuations_as_ints : Array[0.."_SELECT_STATION_BUTTON_COUNT"] of Int;
      actuation_pulses : Array[0.."_SELECT_STATION_BUTTON_COUNT"] of Bool;
      actuation_pulses_as_int : Array[0.."_SELECT_STATION_BUTTON_COUNT"] of Int;
      blank_station : "Station: Single Station";
      i : Int;
      nav_pulses : Int;
      p_stn : DInt;
      selectable_stns_as_dint : Array[0.."STATION_COUNT"] of DInt;
      t_selection_change : "Station Selection Change";
   END_VAR
   // visable_stns[0] := 0;
   // visable_stns[1] := 1;
   // visable_stns[2] := 2;
   // visable_stns[3] := 3;
   // visable_stns[4] := 4;
   // visable_stns[5] := 5;
   // visable_stns[6] := 6;
   // visable_stns[7] := 7;
   // visable_stns[8] := 8;
   // visable_stns[9] := 9;
   // visable_stns[10] := 10;
   // visable_stns[11] := 11;
BEGIN
   REGION "ANIMATIONS"
       "Pop Up: Select Stations: Animations"(all_stations := #all_stations,
                                             meta_data := #meta_data,
                                             visable_stns := #visable_stns,
                                             interface := #interface);
   END_REGION


   REGION "CLEAR SELECTION CHANGE"
       #meta_data.station_selection_change := #t_selection_change;
   END_REGION


   REGION "SELECT STATION BUTTON PULSES"
       "Pop Up: Map Select Button Actuations"(screen_elements := #interface.stn_select_btns,
                                              actuations_as_ints := #actuations_as_ints);
       #"inst Select Station Button Pulses"(btns := #actuations_as_ints,
                                            pulses := #actuation_pulses_as_int);
       "Pop Up: Select Stations: Pulse Ints to Bools"(pulses_as_ints := #actuation_pulses_as_int,
                                                      pulses_as_bools => #actuation_pulses);
   END_REGION


   REGION "PERFORM STATION SELECTION"
       FOR #i := 0 TO "_SELECT_STATION_BUTTON_COUNT" DO
           IF #visable_stns[#i] <> -1 THEN
               "Toggle"(pulse := #actuation_pulses[#i],
                        state := #meta_data.selected_stations.stns[#visable_stns[#i]]);
           END_IF;
       END_FOR;
       #meta_data.selected_stations.count := "Count Selected Stations"(#meta_data.selected_stations.stns);
   END_REGION


   REGION "SCAN FOR CHANGE TO STATION SELECTION"
       #"inst Selection Change"(selected_stns := #meta_data.#selected_stations,
                                station_change => #meta_data.station_selection_change);
   END_REGION


   REGION "BUILD SELECTABLE STATION LIST"
       IF #meta_data.station_selection_change.selection_change OR "FirstScan" THEN
           "Pop Up: Select Stations: Build Selectable Station List"(saved_wips := #saved_WIPs,
                                                                    all_stations := #all_stations,
                                                                    meta_data := #meta_data);
       END_IF;
   END_REGION


   REGION "TABLE NAV"

       // when there are more selectable stations than buttons
       IF #meta_data.selectable_stations.count > "_SELECT_STATION_BUTTON_COUNT" THEN
           #"inst Table Nav"(first_null_index := #meta_data.selectable_stations.count,
                             tblData := #selectable_stns_as_dint,
                             tblDisp := #vis_stns_as_dint,
                             tableNav := #interface.nav_bar.plc,
                             rowIndices := #vis_stns_as_dint);
           // patch for table nav to work with selectable stations
           #"inst Patch for Table Nav in Select Station Popup"(nav_bar := #interface.nav_bar.plc,
                                                               meta_data := #meta_data,
                                                               vis_stns_as_dint := #vis_stns_as_dint,
                                                               visable_stns := #visable_stns);
       END_IF;

       // when there are fewer selectable stations than buttons
       IF #meta_data.selectable_stations.count <= "_SELECT_STATION_BUTTON_COUNT" + 1 THEN
           IF #meta_data.station_selection_change.selection_change THEN
               "Array.Int.Fill"(value:="NULL_TOKEN",
                                int_array := #visable_stns);
               FOR #i := 0 TO #meta_data.selectable_stations.count - 1 DO
                   #visable_stns[#i] := #meta_data.selectable_stations.stns[#i];
               END_FOR;
           END_IF;
       END_IF;


   END_REGION
END_FUNCTION_BLOCK

FUNCTION_BLOCK "Selected_Stations.Selection_Change"   // FB23, SCL
{ S7_Optimized_Access := 'TRUE' }
VERSION : 0.1
   VAR_INPUT
      selected_stns : "Selected Stations";
   END_VAR
   VAR_OUTPUT
      station_change : "Station Selection Change";
   END_VAR
   VAR
      old : Struct
         selected_stns : "Selected Stations";
      END_STRUCT;
   END_VAR
   VAR_TEMP
      i : Int;
      ret : "Station Selection Change";
   END_VAR
BEGIN
   REGION "SCAN FOR CHANGE"
       FOR #i := 0 TO "STATION_COUNT" DO
           IF #selected_stns.stns[#i] <> #old.selected_stns.stns[#i] THEN
               #ret.selection_change := TRUE;
               #ret.station_index := #i;
               IF #selected_stns.stns[#i] AND NOT #old.selected_stns.stns[#i] THEN
                   #ret.rising := TRUE;
                   #ret.falling := FALSE;
               END_IF;
               IF NOT #selected_stns.stns[#i] AND #old.selected_stns.stns[#i] THEN
                   #ret.rising := FALSE;
                   #ret.falling := TRUE;
               END_IF;
               EXIT;
           END_IF;
       END_FOR;
   END_REGION


   REGION "SAVE TO OLD"
       #old.selected_stns := #selected_stns;
   END_REGION


   REGION "RETURN"
       #station_change.falling := #ret.falling;
       #station_change.rising := #ret.rising;
       #station_change.selection_change := #ret.selection_change;
       #station_change.station_index := #ret.station_index;
   END_REGION
END_FUNCTION_BLOCK

FUNCTION_BLOCK "Patch for Table Nav in Select Station Popup"   // FB24, SCL
{ S7_Optimized_Access := 'TRUE' }